// TIA Portal project "Milk_P_2" (V17)

(* hardware
DEVICE "S7-1200 station_1"  S7-1200 Station
   slot 0: "Rack_0"  S7-1200 Rack  Rack  V1.0
   slot 1: "PLC_1"  CPU 1217C DC/DC/DC  6ES7 217-1AG40-0XB0  V4.5
   slot 2: "DI 8x24VDC_1"  6ES7 221-1BF32-0XB0  V2.0
   slot 3: "DQ 8x24VDC _1"  SM 1222 DQ8 x 24VDC  6ES7 222-1BF32-0XB0  V2.0
DEVICE "HMI_1"  KTP700 Basic PN
   slot 0: "HMI_1"  KTP700 Basic PN  6AV2 123-2GB03-0AX0  17.0.0.0
   slot 1: "HMI_RT_1"  KTP700 Basic PN  6AV2 123-2GB03-0AX0  17.0.0.0
   slot 5: "HMI_1.IE_CP_1"  PROFINET Interface  17.0.0.0
      slot 1: "PROFINET Interface_1"  PROFINET Interface
         slot 1: "Port_1"  Port
*)

// ===== PLC "PLC_1"  CPU 1217C DC/DC/DC =====

VAR_GLOBAL   // PLC tag table "Default tag table"
   "Cycle_on_Memory_Bit" AT %M100.0 : Bool;
   "Low_Level_Sensor" AT %M1.0 : Bool;
   "High_Level_Sensor" AT %M1.1 : Bool;
   "Pump_1" AT %Q1.0 : Bool;
   "Milk_Level" AT %MD50 : Real;
   "Start_Fill" AT %M2.0 : Bool;
   "Stop_Fill" AT %M2.1 : Bool;
   "Drain_Start" AT %M2.2 : Bool;
   "Drain_Stop" AT %M2.3 : Bool;
   "Cycle_on_Memory_Bit_2" AT %M200.0 : Bool;
   "Pump_2" AT %Q1.1 : Bool;
   "Sep_Start" AT %M2.4 : Bool;
   "Sep_Stop" AT %M2.5 : Bool;
   "Sep_Memory_Bit" AT %M2.6 : Bool;
   "Clock_Byte" AT %MB0 : Byte;
   "Clock_10Hz" AT %M0.0 : Bool;
   "Clock_5Hz" AT %M0.1 : Bool;
   "Clock_2.5Hz" AT %M0.2 : Bool;
   "Clock_2Hz" AT %M0.3 : Bool;
   "Clock_1.25Hz" AT %M0.4 : Bool;
   "Clock_1Hz" AT %M0.5 : Bool;
   "Clock_0.625Hz" AT %M0.6 : Bool;
   "Clock_0.5Hz" AT %M0.7 : Bool;
   "HMI_Mixer" AT %M2.7 : Bool;
   "Pump_3" AT %Q0.3 : Bool;
   "Furnace_ON" AT %M4.3 : Bool;
   "Furnace_Temp_Sensor" AT %MW4 : Int;
   "Cycle_on_Memory_Bit_3" AT %M50.0 : Bool;
   "Current_Milk_Temp" AT %MW8 : Int;
   "Start_HE" AT %M1.2 : Bool;
   "Stop_HE" AT %M1.3 : Bool;
   "memory_1" AT %M1.4 : Bool;
   "Inıtial_Milk_Temp" AT %MW16 : Int;
   "Wanted_Milk_Temp" AT %MW10 : Int;
   "Heating" AT %Q0.4 : Bool;
   "Cooling_Temp_Sensor" AT %MW12 : Int;
   "Cooling_ON" AT %M1.5 : Bool;
   "Start_CL" AT %M1.6 : Bool;
   "Stop_CL" AT %M1.7 : Bool;
   "Cycle_on_Memory_Bit_4" AT %M7.0 : Bool;
   "memory_2" AT %M7.1 : Bool;
   "Cold_Milk_Temp" AT %MW14 : Int;
   "Heating_OFF" AT %M7.2 : Bool;
   "Cooling_OFF" AT %M7.4 : Bool;
   "Milk_Level_2" AT %MD18 : Real;
   "Low_Level_2" AT %M22.0 : Bool;
   "High_Level_2" AT %M26.0 : Bool;
   "Memory_3" AT %M7.5 : Bool;
   "working" AT %M28.0 : Bool;
   "Start_Package" AT %M28.1 : Bool;
END_VAR

DATA_BLOCK "Bottle Calculation_DB"   // DB1
{ S7_Optimized_Access := 'TRUE' }
VERSION : 0.1
// stored: InstanceOfName Bottle Calculation
"Bottle Calculation"
BEGIN
END_DATA_BLOCK

DATA_BLOCK "Cooling_DB"   // DB2
{ S7_Optimized_Access := 'TRUE' }
VERSION : 0.1
// stored: InstanceOfName Cooling
"Cooling"
BEGIN
END_DATA_BLOCK

DATA_BLOCK "Milk_Pasteurization_DB"   // DB9
{ S7_Optimized_Access := 'TRUE' }
VERSION : 0.1
   VAR
      Fire_Alarm : Bool;
      Warning_Lights : Bool;
      Water_Mist_System : Bool;
   END_VAR
BEGIN
END_DATA_BLOCK

DATA_BLOCK "Heat_Exchange_DB_1"   // DB11
{ S7_Optimized_Access := 'TRUE' }
VERSION : 0.1
// stored: InstanceOfName Heat_Exchange
"Heat_Exchange"
BEGIN
END_DATA_BLOCK

DATA_BLOCK "Pasteurized_Tank_fill_DB"   // DB12
{ S7_Optimized_Access := 'TRUE' }
VERSION : 0.1
// stored: InstanceOfName Pasteurized_Tank_fill
"Pasteurized_Tank_fill"
BEGIN
END_DATA_BLOCK

DATA_BLOCK "Tank_Fill_Drain_DB_1"   // DB13
{ S7_Optimized_Access := 'TRUE' }
VERSION : 0.1
// stored: InstanceOfName Tank_Fill_Drain
"Tank_Fill_Drain"
BEGIN
END_DATA_BLOCK

DATA_BLOCK "Fat_Seperator_DB"   // DB14
{ S7_Optimized_Access := 'TRUE' }
VERSION : 0.1
// stored: InstanceOfName Fat_Seperator
"Fat_Seperator"
BEGIN
END_DATA_BLOCK

// folder: System blocks/Program resources

DATA_BLOCK "Milk_Tank_Timer_1"   // DB3
{ S7_Optimized_Access := 'TRUE' }
AUTHOR : Simatic
FAMILY : IEC
NAME : IEC_TMR
VERSION : 1.0
// stored: InstanceOfName IEC_TIMER
"IEC_TIMER"
BEGIN
END_DATA_BLOCK

DATA_BLOCK "Milk_Tank_Timer_2"   // DB4
{ S7_Optimized_Access := 'TRUE' }
AUTHOR : Simatic
FAMILY : IEC
NAME : IEC_TMR
VERSION : 1.0
// stored: InstanceOfName IEC_TIMER
"IEC_TIMER"
BEGIN
END_DATA_BLOCK

DATA_BLOCK "Sep_Timer"   // DB5
{ S7_Optimized_Access := 'TRUE' }
AUTHOR : Simatic
FAMILY : IEC
NAME : IEC_TMR
VERSION : 1.0
// stored: InstanceOfName IEC_TIMER
"IEC_TIMER"
BEGIN
END_DATA_BLOCK

DATA_BLOCK "HE_Timer1"   // DB6
{ S7_Optimized_Access := 'TRUE' }
AUTHOR : Simatic
FAMILY : IEC
NAME : IEC_TMR
VERSION : 1.0
// stored: InstanceOfName IEC_TIMER
"IEC_TIMER"
BEGIN
END_DATA_BLOCK

DATA_BLOCK "Cooling_Timer"   // DB7
{ S7_Optimized_Access := 'TRUE' }
AUTHOR : Simatic
FAMILY : IEC
NAME : IEC_TMR
VERSION : 1.0
// stored: InstanceOfName IEC_TIMER
"IEC_TIMER"
BEGIN
END_DATA_BLOCK

DATA_BLOCK "P_Tank_Timer1"   // DB8
{ S7_Optimized_Access := 'TRUE' }
AUTHOR : Simatic
FAMILY : IEC
NAME : IEC_TMR
VERSION : 1.0
// stored: InstanceOfName IEC_TIMER
"IEC_TIMER"
BEGIN
END_DATA_BLOCK

DATA_BLOCK "Bottle Counter"   // DB10
{ S7_Optimized_Access := 'TRUE' }
AUTHOR : Simatic
FAMILY : IEC
NAME : CNTR
VERSION : 1.0
// stored: InstanceOfName IEC_COUNTER
"IEC_COUNTER"
BEGIN
END_DATA_BLOCK

// folder: (top level)

FUNCTION_BLOCK "Tank_Fill_Drain"   // FB1, LAD
{ S7_Optimized_Access := 'TRUE' }
VERSION : 0.1
   VAR_INPUT
      "Fill Start" : Bool;
      "Fill Stop" : Bool;
      "Drain Start" : Bool;
      "Drain Stop" : Bool;
   END_VAR
   VAR_OUTPUT
      "Milk Level" : Real;
      "Low Level" : Bool;
      "Pump 2" : Bool;
      Pump : Bool;
      "High Level" : Bool;
   END_VAR
   VAR
      Inıtial_Fat_P : Real := 4.0;
   END_VAR
   VAR_TEMP
      Fat_temp : Real;
   END_VAR
   VAR_TEMP   // added for the SCL form of the ladder/FBD networks
      _w1 : Bool;
   END_VAR
BEGIN

REGION Network 1: Start_Fill System
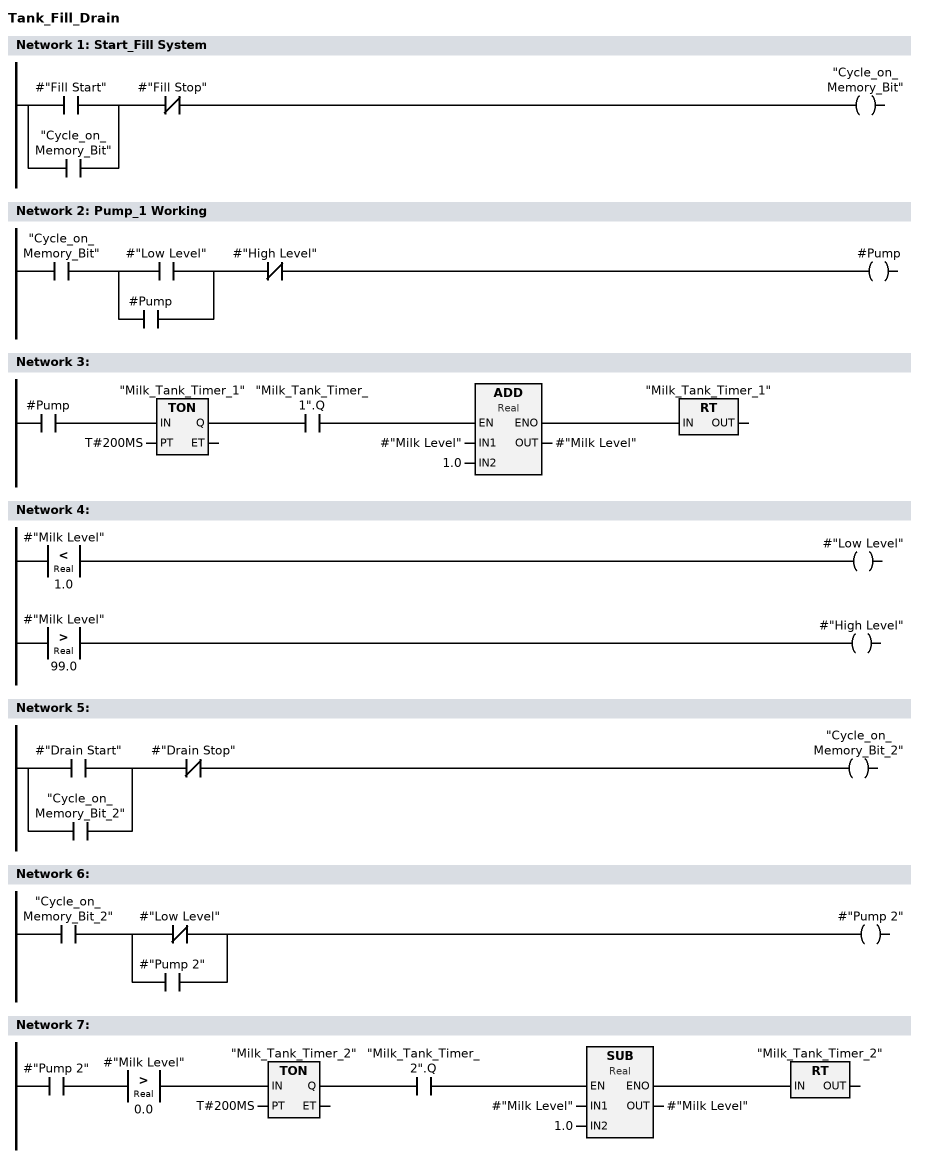
   RUNG wire#powerrail
      Contact( #"Fill Start" )
      wire#w1
      I_Contact( #"Fill Stop" )
      Coil( "Cycle_on_Memory_Bit" )
   END_RUNG
   RUNG wire#powerrail
      Contact( "Cycle_on_Memory_Bit" )
   END_RUNG wire#w1
   // the same network as SCL:
   "Cycle_on_Memory_Bit" := (#"Fill Start" OR "Cycle_on_Memory_Bit") AND NOT #"Fill Stop";
END_REGION

REGION Network 2: Pump_1 Working
   RUNG wire#powerrail
      Contact( "Cycle_on_Memory_Bit" )
      wire#w1
      Contact( #"Low Level" )
      wire#w2
      I_Contact( #"High Level" )
      Coil( #Pump )
   END_RUNG
   RUNG wire#w1
      Contact( #Pump )
   END_RUNG wire#w2
   // the same network as SCL:
   #Pump := "Cycle_on_Memory_Bit" AND (#"Low Level" OR #Pump) AND NOT #"High Level";
END_REGION

REGION Network 3
   "Milk_Tank_Timer_1".TON(IN := #Pump, PT := T#200MS);
   #_w1 := "Milk_Tank_Timer_1".Q AND "Milk_Tank_Timer_1".Q;
   IF #_w1 THEN
       #"Milk Level" := #"Milk Level" + 1.0;
       RESET_TIMER("Milk_Tank_Timer_1");
   END_IF;
END_REGION

REGION Network 4
   RUNG wire#powerrail
      { S7_Templates := "SrcType := Real" } LT_Contact(in1 := #"Milk Level", in2 := 1.0)
      Coil( #"Low Level" )
   END_RUNG
   RUNG wire#powerrail
      { S7_Templates := "SrcType := Real" } GT_Contact(in1 := #"Milk Level", in2 := 99.0)
      Coil( #"High Level" )
   END_RUNG
   // the same network as SCL:
   #"Low Level" := #"Milk Level" < 1.0;
   #"High Level" := #"Milk Level" > 99.0;
END_REGION

REGION Network 5
   RUNG wire#powerrail
      Contact( #"Drain Start" )
      wire#w1
      I_Contact( #"Drain Stop" )
      Coil( "Cycle_on_Memory_Bit_2" )
   END_RUNG
   RUNG wire#powerrail
      Contact( "Cycle_on_Memory_Bit_2" )
   END_RUNG wire#w1
   // the same network as SCL:
   "Cycle_on_Memory_Bit_2" := (#"Drain Start" OR "Cycle_on_Memory_Bit_2") AND NOT #"Drain Stop";
END_REGION

REGION Network 6
   RUNG wire#powerrail
      Contact( "Cycle_on_Memory_Bit_2" )
      wire#w1
      I_Contact( #"Low Level" )
      wire#w2
      Coil( #"Pump 2" )
   END_RUNG
   RUNG wire#w1
      Contact( #"Pump 2" )
   END_RUNG wire#w2
   // the same network as SCL:
   #"Pump 2" := "Cycle_on_Memory_Bit_2" AND (NOT #"Low Level" OR #"Pump 2");
END_REGION

REGION Network 7
   "Milk_Tank_Timer_2".TON(IN := #"Pump 2" AND (#"Milk Level" > 0.0), PT := T#200MS);
   #_w1 := "Milk_Tank_Timer_2".Q AND "Milk_Tank_Timer_2".Q;
   IF #_w1 THEN
       #"Milk Level" := #"Milk Level" - 1.0;
       RESET_TIMER("Milk_Tank_Timer_2");
   END_IF;
END_REGION
END_FUNCTION_BLOCK

FUNCTION_BLOCK "Heat_Exchange"   // FB2, LAD
{ S7_Optimized_Access := 'TRUE' }
VERSION : 0.1
   VAR_INPUT
      "Heat Exchanger Start" : Bool;
      "Heat Exchanger Stop" : Bool;
   END_VAR
   VAR_OUTPUT
      "Furnace ON" : Bool;
      "Current Milk Temperature" : Int;
   END_VAR
   VAR
      heat_difference : Int;
      addition_step : Int;
      furnace_temp_sensor : Int := 500;
      "wanted milk temp" : Int := 72;
      "Initial Temperature" : Int := 20;
   END_VAR
   VAR_TEMP   // added for the SCL form of the ladder/FBD networks
      _w1 : Bool;
   END_VAR
BEGIN

REGION Network 1
   // While loop
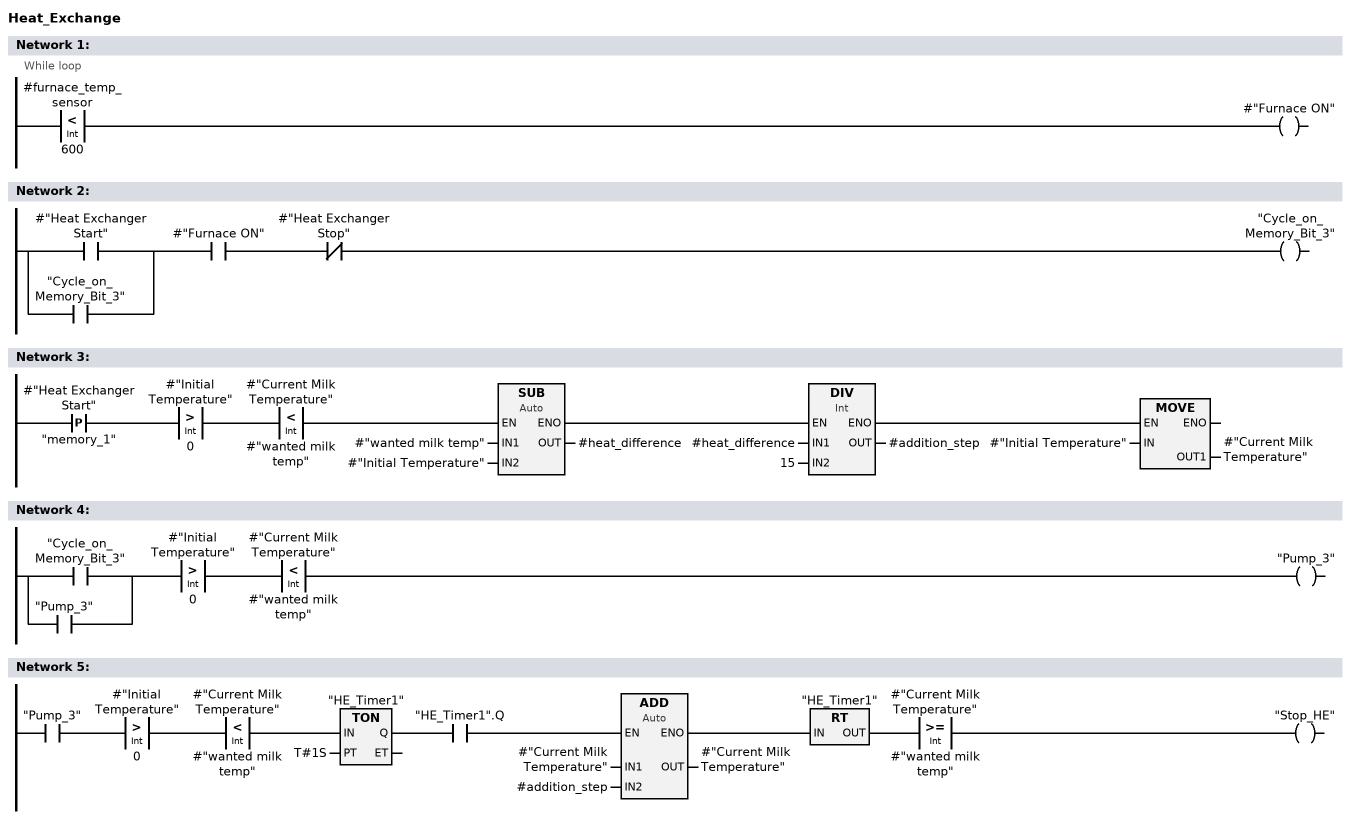
   RUNG wire#powerrail
      { S7_Templates := "SrcType := Int" } LT_Contact(in1 := #furnace_temp_sensor, in2 := 600)
      Coil( #"Furnace ON" )
   END_RUNG
   // the same network as SCL:
   #"Furnace ON" := #furnace_temp_sensor < 600;
END_REGION

REGION Network 2
   RUNG wire#powerrail
      Contact( #"Heat Exchanger Start" )
      wire#w1
      Contact( #"Furnace ON" )
      I_Contact( #"Heat Exchanger Stop" )
      Coil( "Cycle_on_Memory_Bit_3" )
   END_RUNG
   RUNG wire#powerrail
      Contact( "Cycle_on_Memory_Bit_3" )
   END_RUNG wire#w1
   // the same network as SCL:
   "Cycle_on_Memory_Bit_3" := (#"Heat Exchanger Start" OR "Cycle_on_Memory_Bit_3") AND #"Furnace ON" AND NOT #"Heat Exchanger Stop";
END_REGION

REGION Network 3
   RUNG wire#powerrail
      P_Contact(operand := #"Heat Exchanger Start", bit := "memory_1")
      { S7_Templates := "SrcType := Int" } GT_Contact(in1 := #"Initial Temperature", in2 := 0)
      { S7_Templates := "SrcType := Int" } LT_Contact(in1 := #"Current Milk Temperature", in2 := #"wanted milk temp")
      Sub(in1 := #"wanted milk temp", in2 := #"Initial Temperature", out => #heat_difference)
      { S7_Templates := "SrcType := Int" } Div(in1 := #heat_difference, in2 := 15, out => #addition_step)
      Move(in := #"Initial Temperature", out1 => #"Current Milk Temperature")
   END_RUNG
   // the same network as SCL:
   #_w1 := #"Heat Exchanger Start" AND NOT "memory_1";   // rising edge of #"Heat Exchanger Start"
   "memory_1" := #"Heat Exchanger Start";
   IF #_w1 AND (#"Initial Temperature" > 0) AND (#"Current Milk Temperature" < #"wanted milk temp") THEN
       #heat_difference := #"wanted milk temp" - #"Initial Temperature";
       #addition_step := #heat_difference / 15;
       #"Current Milk Temperature" := #"Initial Temperature";
   END_IF;
END_REGION

REGION Network 4
   RUNG wire#powerrail
      Contact( "Cycle_on_Memory_Bit_3" )
      wire#w1
      { S7_Templates := "SrcType := Int" } GT_Contact(in1 := #"Initial Temperature", in2 := 0)
      { S7_Templates := "SrcType := Int" } LT_Contact(in1 := #"Current Milk Temperature", in2 := #"wanted milk temp")
      Coil( "Pump_3" )
   END_RUNG
   RUNG wire#powerrail
      Contact( "Pump_3" )
   END_RUNG wire#w1
   // the same network as SCL:
   "Pump_3" := ("Cycle_on_Memory_Bit_3" OR "Pump_3") AND (#"Initial Temperature" > 0) AND (#"Current Milk Temperature" < #"wanted milk temp");
END_REGION

REGION Network 5
   "HE_Timer1".TON(IN := "Pump_3" AND (#"Initial Temperature" > 0) AND (#"Current Milk Temperature" < #"wanted milk temp"),
                   PT := T#1S);
   #_w1 := "HE_Timer1".Q AND "HE_Timer1".Q;
   IF #_w1 THEN
       #"Current Milk Temperature" := #"Current Milk Temperature" + #addition_step;
       RESET_TIMER("HE_Timer1");
   END_IF;
   "Stop_HE" := #_w1 AND (#"Current Milk Temperature" >= #"wanted milk temp");
END_REGION
END_FUNCTION_BLOCK

FUNCTION_BLOCK "Cooling"   // FB3, LAD
{ S7_Optimized_Access := 'TRUE' }
VERSION : 0.1
   VAR_OUTPUT
      "Cooling OFF" : Bool;
      "Cooling ON" : Bool;
   END_VAR
   VAR
      heat_diff : Int;
      diff_step : Int;
      Wanted_cold_milk : Int := 4;
      "Current Temp" : Int;
      cooling_temp_sensor : Int := -15;
   END_VAR
   VAR_TEMP   // added for the SCL form of the ladder/FBD networks
      _w1 : Bool;
   END_VAR
BEGIN

REGION Network 1
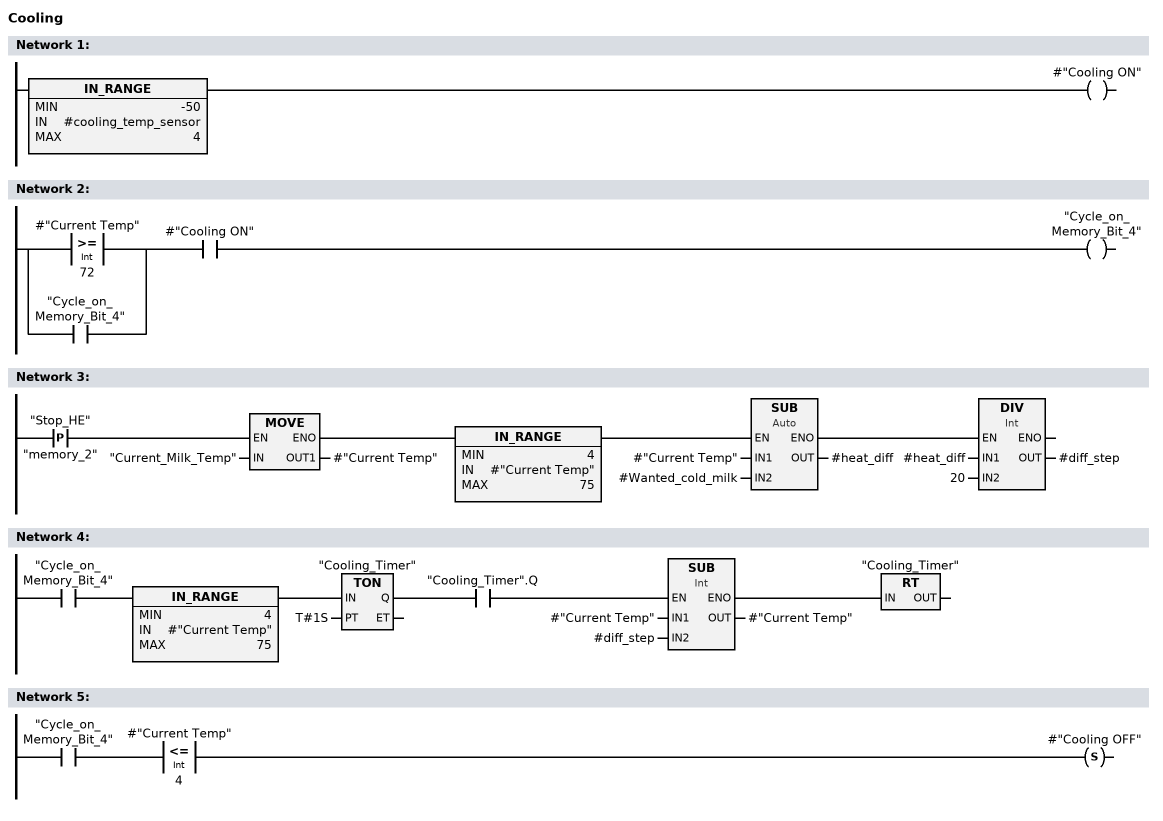
   RUNG wire#powerrail
      { S7_Templates := "SrcType := Int" } InRange(min := -50, in := #cooling_temp_sensor, max := 4)
      Coil( #"Cooling ON" )
   END_RUNG
   // the same network as SCL:
   #"Cooling ON" := (-50 <= #cooling_temp_sensor) AND (#cooling_temp_sensor <= 4);
END_REGION

REGION Network 2
   RUNG wire#powerrail
      { S7_Templates := "SrcType := Int" } GE_Contact(in1 := #"Current Temp", in2 := 72)
      wire#w1
      Contact( #"Cooling ON" )
      Coil( "Cycle_on_Memory_Bit_4" )
   END_RUNG
   RUNG wire#powerrail
      Contact( "Cycle_on_Memory_Bit_4" )
   END_RUNG wire#w1
   // the same network as SCL:
   "Cycle_on_Memory_Bit_4" := ((#"Current Temp" >= 72) OR "Cycle_on_Memory_Bit_4") AND #"Cooling ON";
END_REGION

REGION Network 3
   RUNG wire#powerrail
      P_Contact(operand := "Stop_HE", bit := "memory_2")
      Move(in := "Current_Milk_Temp", out1 => #"Current Temp")
      { S7_Templates := "SrcType := Int" } InRange(min := 4, in := #"Current Temp", max := 75)
      Sub(in1 := #"Current Temp", in2 := #Wanted_cold_milk, out => #heat_diff)
      { S7_Templates := "SrcType := Int" } Div(in1 := #heat_diff, in2 := 20, out => #diff_step)
   END_RUNG
   // the same network as SCL:
   #_w1 := "Stop_HE" AND NOT "memory_2";   // rising edge of "Stop_HE"
   "memory_2" := "Stop_HE";
   IF #_w1 THEN #"Current Temp" := "Current_Milk_Temp"; END_IF;
   IF #_w1 AND (4 <= #"Current Temp") AND (#"Current Temp" <= 75) THEN
       #heat_diff := #"Current Temp" - #Wanted_cold_milk;
       #diff_step := #heat_diff / 20;
   END_IF;
END_REGION

REGION Network 4
   "Cooling_Timer".TON(IN := "Cycle_on_Memory_Bit_4" AND (4 <= #"Current Temp") AND (#"Current Temp" <= 75),
                       PT := T#1S);
   #_w1 := "Cooling_Timer".Q AND "Cooling_Timer".Q;
   IF #_w1 THEN
       #"Current Temp" := #"Current Temp" - #diff_step;
       RESET_TIMER("Cooling_Timer");
   END_IF;
END_REGION

REGION Network 5
   RUNG wire#powerrail
      Contact( "Cycle_on_Memory_Bit_4" )
      { S7_Templates := "SrcType := Int" } LE_Contact(in1 := #"Current Temp", in2 := 4)
      S_Coil( #"Cooling OFF" )
   END_RUNG
   // the same network as SCL:
   IF "Cycle_on_Memory_Bit_4" AND (#"Current Temp" <= 4) THEN #"Cooling OFF" := TRUE; END_IF;
END_REGION
END_FUNCTION_BLOCK

FUNCTION_BLOCK "Fat_Seperator"   // FB4, LAD
{ S7_Optimized_Access := 'TRUE' }
VERSION : 0.1
   VAR_INPUT
      "Seperator Start" : Bool;
      "Seperator Stop" : Bool;
   END_VAR
   VAR_OUTPUT
      "Fat Percantage" : Int := 4;
   END_VAR
   VAR
      wanted_fat : Int := 2;
      diff : Int;
   END_VAR
BEGIN

REGION Network 1
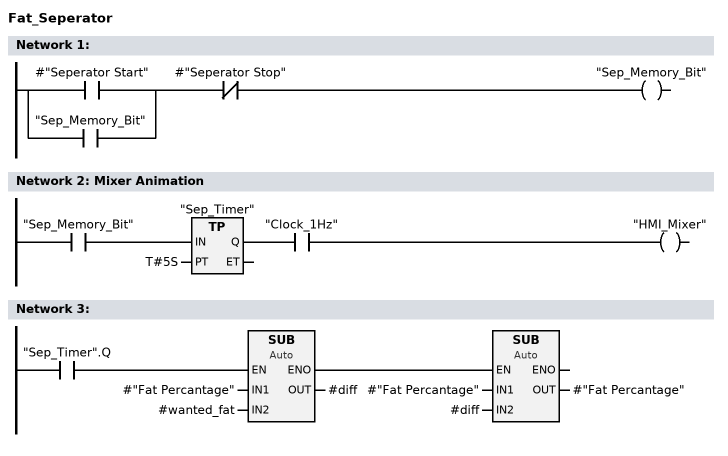
   RUNG wire#powerrail
      Contact( #"Seperator Start" )
      wire#w1
      I_Contact( #"Seperator Stop" )
      Coil( "Sep_Memory_Bit" )
   END_RUNG
   RUNG wire#powerrail
      Contact( "Sep_Memory_Bit" )
   END_RUNG wire#w1
   // the same network as SCL:
   "Sep_Memory_Bit" := (#"Seperator Start" OR "Sep_Memory_Bit") AND NOT #"Seperator Stop";
END_REGION

REGION Network 2: Mixer Animation
   "Sep_Timer".TP(IN := "Sep_Memory_Bit", PT := T#5S);
   "HMI_Mixer" := "Sep_Timer".Q AND "Clock_1Hz";
END_REGION

REGION Network 3
   RUNG wire#powerrail
      Contact( "Sep_Timer".Q )
      Sub(in1 := #"Fat Percantage", in2 := #wanted_fat, out => #diff)
      Sub(in1 := #"Fat Percantage", in2 := #diff, out => #"Fat Percantage")
   END_RUNG
   // the same network as SCL:
   IF "Sep_Timer".Q THEN
       #diff := #"Fat Percantage" - #wanted_fat;
       #"Fat Percantage" := #"Fat Percantage" - #diff;
   END_IF;
END_REGION
END_FUNCTION_BLOCK

FUNCTION_BLOCK "Pasteurized_Tank_fill"   // FB5, LAD
{ S7_Optimized_Access := 'TRUE' }
VERSION : 0.1
   VAR_INPUT
      Start : Bool;
      Stop : Bool;
   END_VAR
   VAR_OUTPUT
      low : Bool;
      high : Bool;
      working : Bool;
      milk_level : Real;
   END_VAR
   VAR_TEMP   // added for the SCL form of the ladder/FBD networks
      _w1 : Bool;
   END_VAR
BEGIN

REGION Network 1
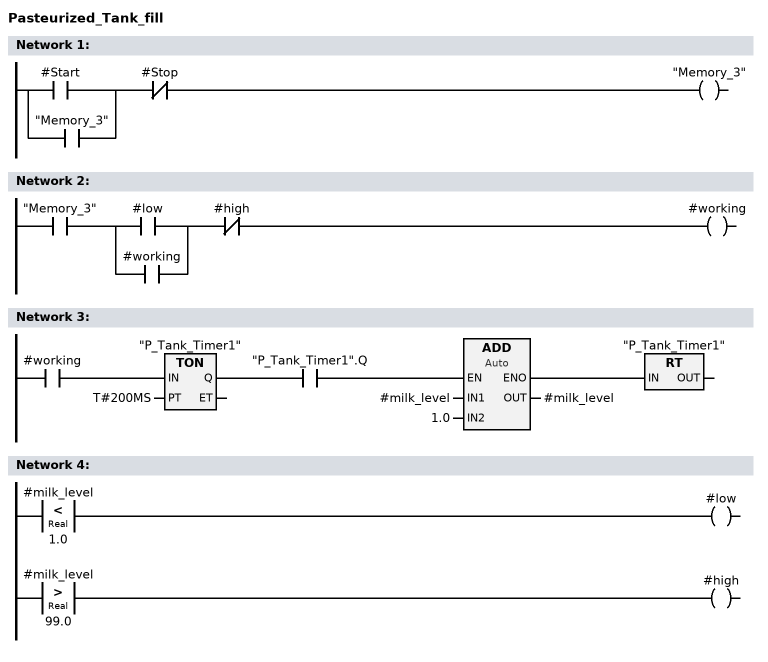
   RUNG wire#powerrail
      Contact( #Start )
      wire#w1
      I_Contact( #Stop )
      Coil( "Memory_3" )
   END_RUNG
   RUNG wire#powerrail
      Contact( "Memory_3" )
   END_RUNG wire#w1
   // the same network as SCL:
   "Memory_3" := (#Start OR "Memory_3") AND NOT #Stop;
END_REGION

REGION Network 2
   RUNG wire#powerrail
      Contact( "Memory_3" )
      wire#w1
      Contact( #low )
      wire#w2
      I_Contact( #high )
      Coil( #working )
   END_RUNG
   RUNG wire#w1
      Contact( #working )
   END_RUNG wire#w2
   // the same network as SCL:
   #working := "Memory_3" AND (#low OR #working) AND NOT #high;
END_REGION

REGION Network 3
   "P_Tank_Timer1".TON(IN := #working, PT := T#200MS);
   #_w1 := "P_Tank_Timer1".Q AND "P_Tank_Timer1".Q;
   IF #_w1 THEN
       #milk_level := #milk_level + 1.0;
       RESET_TIMER("P_Tank_Timer1");
   END_IF;
END_REGION

REGION Network 4
   RUNG wire#powerrail
      { S7_Templates := "SrcType := Real" } LT_Contact(in1 := #milk_level, in2 := 1.0)
      Coil( #low )
   END_RUNG
   RUNG wire#powerrail
      { S7_Templates := "SrcType := Real" } GT_Contact(in1 := #milk_level, in2 := 99.0)
      Coil( #high )
   END_RUNG
   // the same network as SCL:
   #low := #milk_level < 1.0;
   #high := #milk_level > 99.0;
END_REGION
END_FUNCTION_BLOCK

FUNCTION_BLOCK "Bottle Calculation"   // FB6, LAD
{ S7_Optimized_Access := 'TRUE' }
VERSION : 0.1
   VAR_INPUT
      "Start Packaging" : Bool;
   END_VAR
   VAR_OUTPUT
      "Bottle Count" : Int;
   END_VAR
   VAR
      C1 : Bool;
      "Milk Litres" : Real := 10.0;
      "Bottle Litres" : Real := 0.35;
      Running : Bool;
   END_VAR
   VAR_TEMP   // added for the SCL form of the ladder/FBD networks
      _w1 : Bool;
   END_VAR
BEGIN

REGION Network 1
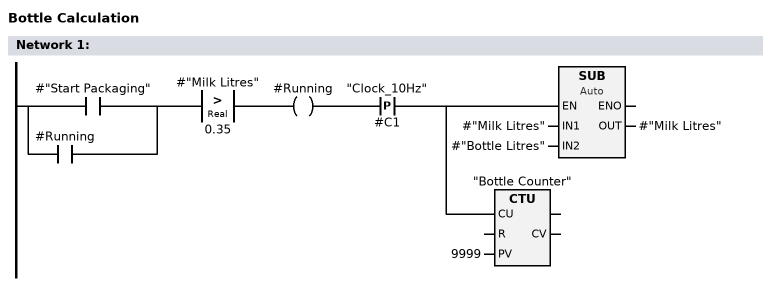
   #Running := (#"Start Packaging" OR #Running) AND (#"Milk Litres" > 0.35);
   #_w1 := #Running AND "Clock_10Hz" AND NOT #C1;   // rising edge of "Clock_10Hz"
   #C1 := "Clock_10Hz";
   IF #_w1 THEN #"Milk Litres" := #"Milk Litres" - #"Bottle Litres"; END_IF;
   "Bottle Counter".CTU(CU := #_w1, PV := 9999);
END_REGION
END_FUNCTION_BLOCK

ORGANIZATION_BLOCK "Main"   // OB1, LAD, ProgramCycle
TITLE = "Main Program Sweep (Cycle)"
{ S7_Optimized_Access := 'TRUE' }
VERSION : 0.1
   VAR_INPUT
      Initial_Call : Bool;   // Initial call of this OB
      Remanence : Bool;   // =True, if remanent data are available
   END_VAR
BEGIN

REGION Network 1: Raw Milk Fill and Drain System
   // Raw milk is filled to a storage tank and it is drain to a fat seperator system.
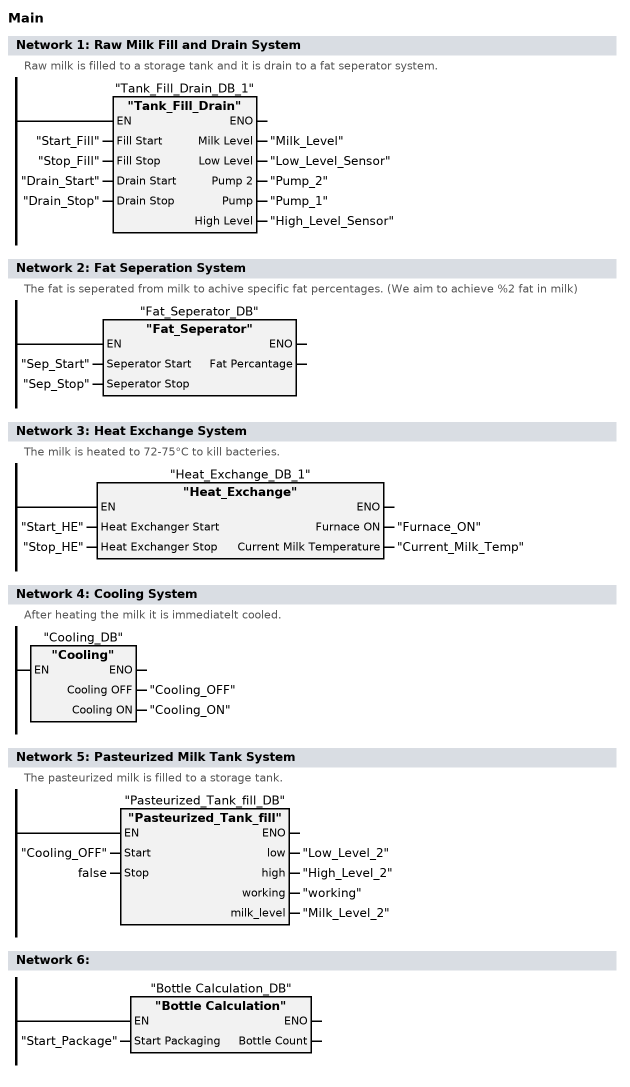
   RUNG wire#powerrail
      "Tank_Fill_Drain_DB_1"("Fill Start" := "Start_Fill", "Fill Stop" := "Stop_Fill", "Drain Start" := "Drain_Start", "Drain Stop" := "Drain_Stop", "Milk Level" => "Milk_Level", "Low Level" => "Low_Level_Sensor", "Pump 2" => "Pump_2", Pump => "Pump_1", "High Level" => "High_Level_Sensor")
   END_RUNG
   // the same network as SCL:
   "Tank_Fill_Drain_DB_1"("Fill Start" := "Start_Fill",   // "Tank_Fill_Drain"
                          "Fill Stop" := "Stop_Fill",
                          "Drain Start" := "Drain_Start",
                          "Drain Stop" := "Drain_Stop",
                          "Milk Level" => "Milk_Level",
                          "Low Level" => "Low_Level_Sensor",
                          "Pump 2" => "Pump_2",
                          Pump => "Pump_1",
                          "High Level" => "High_Level_Sensor");
END_REGION

REGION Network 2: Fat Seperation System
   // The fat is seperated from milk to achive specific fat percentages. (We aim to achieve %2 fat in milk)
   RUNG wire#powerrail
      "Fat_Seperator_DB"("Seperator Start" := "Sep_Start", "Seperator Stop" := "Sep_Stop", "Fat Percantage" =>)
   END_RUNG
   // the same network as SCL:
   "Fat_Seperator_DB"("Seperator Start" := "Sep_Start", "Seperator Stop" := "Sep_Stop");   // "Fat_Seperator"
END_REGION

REGION Network 3: Heat Exchange System
   // The milk is heated to 72-75°C to kill bacteries.
   RUNG wire#powerrail
      "Heat_Exchange_DB_1"("Heat Exchanger Start" := "Start_HE", "Heat Exchanger Stop" := "Stop_HE", "Furnace ON" => "Furnace_ON", "Current Milk Temperature" => "Current_Milk_Temp")
   END_RUNG
   // the same network as SCL:
   "Heat_Exchange_DB_1"("Heat Exchanger Start" := "Start_HE",   // "Heat_Exchange"
                        "Heat Exchanger Stop" := "Stop_HE",
                        "Furnace ON" => "Furnace_ON",
                        "Current Milk Temperature" => "Current_Milk_Temp");
END_REGION

REGION Network 4: Cooling System
   // After heating the milk it is immediatelt cooled.
   RUNG wire#powerrail
      "Cooling_DB"("Cooling OFF" => "Cooling_OFF", "Cooling ON" => "Cooling_ON")
   END_RUNG
   // the same network as SCL:
   "Cooling_DB"("Cooling OFF" => "Cooling_OFF", "Cooling ON" => "Cooling_ON");   // "Cooling"
END_REGION

REGION Network 5: Pasteurized Milk Tank System
   // The pasteurized milk is filled to a storage tank.
   RUNG wire#powerrail
      "Pasteurized_Tank_fill_DB"(Start := "Cooling_OFF", Stop := false, low => "Low_Level_2", high => "High_Level_2", working => "working", milk_level => "Milk_Level_2")
   END_RUNG
   // the same network as SCL:
   "Pasteurized_Tank_fill_DB"(Start := "Cooling_OFF",   // "Pasteurized_Tank_fill"
                           Stop := false,
                           low => "Low_Level_2",
                           high => "High_Level_2",
                           working => "working",
                           milk_level => "Milk_Level_2");
END_REGION

REGION Network 6
   RUNG wire#powerrail
      "Bottle Calculation_DB"("Start Packaging" := "Start_Package", "Bottle Count" =>)
   END_RUNG
   // the same network as SCL:
   "Bottle Calculation_DB"("Start Packaging" := "Start_Package");   // "Bottle Calculation"
END_REGION
END_ORGANIZATION_BLOCK

ORGANIZATION_BLOCK "Cyclic interrupt (HE_FIRE)"   // OB30, LAD, CyclicInterrupt
{ S7_Optimized_Access := 'TRUE' }
VERSION : 0.1
   VAR_INPUT
      Initial_Call : Bool;   // Initial call of this OB
      Event_Count : Int;   // Events discarded
   END_VAR
BEGIN

REGION Network 1
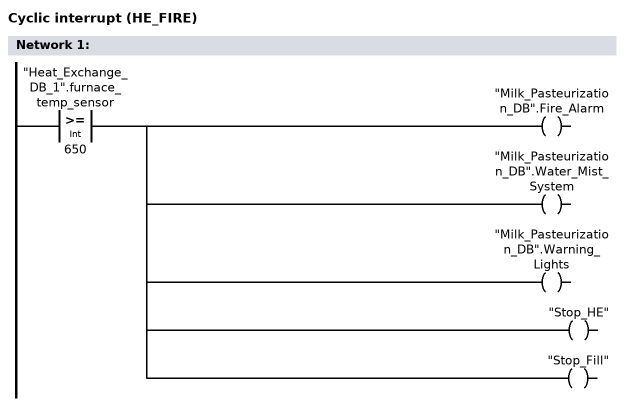
   RUNG wire#powerrail
      { S7_Templates := "SrcType := Int" } GE_Contact(in1 := "Heat_Exchange_DB_1".furnace_temp_sensor, in2 := 650)
      wire#w1
      Coil( "Milk_Pasteurization_DB".Fire_Alarm )
   END_RUNG
   RUNG wire#w1
      Coil( "Milk_Pasteurization_DB".Water_Mist_System )
   END_RUNG
   RUNG wire#w1
      Coil( "Milk_Pasteurization_DB".Warning_Lights )
   END_RUNG
   RUNG wire#w1
      Coil( "Stop_HE" )
   END_RUNG
   RUNG wire#w1
      Coil( "Stop_Fill" )
   END_RUNG
   // the same network as SCL:
   "Milk_Pasteurization_DB".Fire_Alarm := "Heat_Exchange_DB_1".furnace_temp_sensor >= 650;
   "Milk_Pasteurization_DB".Water_Mist_System := "Milk_Pasteurization_DB".Fire_Alarm;
   "Milk_Pasteurization_DB".Warning_Lights := "Milk_Pasteurization_DB".Fire_Alarm;
   "Stop_HE" := "Milk_Pasteurization_DB".Fire_Alarm;
   "Stop_Fill" := "Milk_Pasteurization_DB".Fire_Alarm;
END_REGION
END_ORGANIZATION_BLOCK

(* ===== HMI "HMI_RT_1" =====
system functions are stored by id; their names below are inferred from use
connection "HMI_Connection_1": ETHERNET, SMART_S7_1200_OMS

HMI tags "Default tag table"
   "Tag_ScreenNumber" : UInt, internal
   "Low_Level_Sensor" : Bool = PLC Low_Level_Sensor AT %M1.0, 1 s
   "High_Level_Sensor" : Bool = PLC High_Level_Sensor AT %M1.1, 1 s
   "Water_Level" : Real = PLC Milk_Level AT %MD50, 1 s
   "Start_HMI" : Bool = PLC Start_Fill AT %M2.0, 1 s
   "Stop_HMI" : Bool = PLC Stop_Fill AT %M2.1, 1 s
   "Drain_Start" : Bool = PLC Drain_Start AT %M2.2, 1 s
   "Drain_Stop" : Bool = PLC Drain_Stop AT %M2.3, 1 s
   "Sep_Start" : Bool = PLC Sep_Start AT %M2.4, 100 ms
   "Sep_Stop" : Bool = PLC Sep_Stop AT %M2.5, 100 ms
   "HMI_Mixer" : Bool = PLC HMI_Mixer AT %M2.7, 100 ms
   "Pump_1" : Bool = PLC Pump_1 AT %Q1.0, 100 ms
   "Pump_2" : Bool = PLC Pump_2 AT %Q1.1, 100 ms
   "Start_HE" : Bool = PLC Start_HE AT %M1.2, 1 s
   "Stop_HE" : Bool = PLC Stop_HE AT %M1.3, 1 s
   "Inıtial_Milk_Temp" : Int = PLC Inıtial_Milk_Temp AT %MW16, 1 s
   "Current_Milk_Temp" : Int = PLC Current_Milk_Temp AT %MW8, 1 s
   "Furnace_Temp_Sensor" : Int = PLC Furnace_Temp_Sensor AT %MW4, 1 s
   "Wanted_Milk_Temp" : Int = PLC Wanted_Milk_Temp AT %MW10, 1 s
   "Clock_0.5Hz" : Bool = PLC "Clock_0.5Hz" AT %M0.7, 1 s
   "Clock_10Hz" : Bool = PLC Clock_10Hz AT %M0.0, 1 s
   "Start_CL" : Bool = PLC Start_CL AT %M1.6, 1 s
   "Stop_CL" : Bool = PLC Stop_CL AT %M1.7, 1 s
   "Cold_Milk_Temp" : Int = PLC Cold_Milk_Temp AT %MW14, 1 s
   "Heat_Exchange_DB_1_Initial Temperature" : Int = PLC Heat_Exchange_DB_1."Initial Temperature", 1 s
   "Heat_Exchange_DB_1_wanted milk temp" : Int = PLC Heat_Exchange_DB_1."wanted milk temp", 1 s
   "Heat_Exchange_DB_1_furnace_temp_sensor" : Int = PLC Heat_Exchange_DB_1.furnace_temp_sensor, 1 s
   "Cooling_DB_Wanted_cold_milk" : Int = PLC Cooling_DB.Wanted_cold_milk, 1 s
   "Cooling_DB_Current Temp" : Int = PLC Cooling_DB."Current Temp", 1 s
   "Milk_Level_2" : Real = PLC Milk_Level_2 AT %MD18, 1 s
   "Fat_Seperator_DB_Initial Fat Percantage" : Int = PLC Fat_Seperator_DB."Fat Percantage", 1 s
   "Fat_Seperator_DB_diff" : Int = PLC Fat_Seperator_DB.diff, 1 s
   "Bottle Calculation_DB_Bottle Count" : Int = PLC "Bottle Calculation_DB"."Bottle Count", 1 s
   "Start_Package" : Bool = PLC Start_Package AT %M28.1, 1 s
   "Bottle Counter_CV" : Int = PLC "Bottle Counter".CV, 1 s
   "Low_Level_2" : Bool = PLC Low_Level_2 AT %M22.0, 1 s
   "High_Level_2" : Bool = PLC High_Level_2 AT %M26.0, 1 s

HMI tags "User"
   "Esra Cesur" : WString[254], internal

screen "Root screen" 800x480, template "Template_1"
   on GenerateScreen: SetTag("Stop_HMI", 1)
   Softkey "Softkey_F1" at 0,0 size 0x0
      on KeyDown: ActivateScreen("Root screen", 0)
   Button "Button_3" at 320,349 size 156x119; TextOff 'Cooling'; Authorization "Operator"
      on Click: ActivateScreen("Cooling", 0)
   Button "Button_4" at 479,349 size 156x119; TextOff 'Pasteurized Milk'; Authorization "Operator"
      on Click: ActivateScreen("Pasteurized_Milk", 0)
   Button "Button_5" at 638,349 size 156x119; TextOff 'Log OFF'
      on Click: function_f23ef4c9()
   GraphicView "Graphic view_1" at 0,112 size 800x237; Picture "1009-10099800_cow-milk-cattle"
   Button "Button_2" at 0,349 size 154x119; TextOff 'Raw Milk Tank'; TextOn 'Raw_Milk_Tank'; Authorization "Operator"
      on Click: ActivateScreen("Raw_Milk_Tank", 0)
   Button "Button_1" at 157,349 size 160x119; TextOff 'Heat Exchange'; TextOn 'Heat_Exchange'; Authorization "Operator"
      on Click: ActivateScreen("Heat_Exchange", 0)
   Softkey "Softkey_F8" at 0,0 size 0x0
      on KeyDown: function_f23ef4c9(); ActivateScreen("Root screen", 0)

screen "Raw_Milk_Tank" 800x480
   Softkey "Softkey_F2" at 0,0 size 0x0
      on KeyDown: ActivateScreen("Raw_Milk_Tank", 0)
   Softkey "Softkey_F1" at 0,0 size 0x0
      on KeyDown: ActivateScreen("Root screen", 0)
   GraphicView "Graphic view_19" at 647,214 size 65x49; Picture "Graphic_8"
   GraphicView "Graphic view_18" at 560,291 size 55x48; Picture "Graphic_46"
   GraphicView "Graphic view_10" at 513,97 size 147x222; Picture "Graphic_28"
   GraphicView "Graphic view_12" at 529,133 size 116x119; Picture "Graphic_33"
      Visibility <- "HMI_Mixer"
   GraphicView "Graphic view_11" at 547,126 size 78x94; Picture "Graphic_32"
      Visibility <- "HMI_Mixer"
   GraphicView "Graphic view_20" at 529,133 size 116x119; Picture "Graphic_47"
      Visibility <- "HMI_Mixer"
   GraphicView "Graphic view_21" at 547,126 size 78x94; Picture "Graphic_48"
      Visibility <- "HMI_Mixer"
   GraphicView "Graphic view_23" at 760,215 size 40x51; Picture "Graphic_8"
   GraphicView "Graphic view_17" at 465,140 size 59x47; Picture "Graphic_8"
   GraphicView "Graphic view_7" at 219,338 size 78x57; Picture "Graphic_8"
   GraphicView "Graphic view_3" at 166,340 size 59x53; Picture "Graphic_4"
   GraphicView "Graphic view_1" at 121,113 size 145x239; Picture "Graphic_1"
   Bar "Bar_1" at 138,158 size 112x141; MinimumValue 0; MaximumValue 100
      ProcessValue <- "Water_Level"
   GraphicView "Graphic view_2" at 166,66 size 59x53; Picture "Graphic_3"
   GraphicView "Graphic view_6" at 121,66 size 48x53; Picture "Graphic_8"
   Button "Button_1" at 21,150 size 99x38; TextOff 'Fill Start'
      on Press: function_b14e0dd5("Start_HMI", 0)
      Appearance <- "Start_HMI"
   Button "Button_2" at 21,195 size 100x38; TextOff 'Fill Stop'
      on Press: function_b14e0dd5("Stop_HMI", 0)
      Appearance <- "Stop_HMI"
   Rectangle "Rectangle_1" at 266,253 size 98x22
      Appearance <- "Low_Level_Sensor"
   TextField "Text field_1" at 270,251 size 86x23; Text 'Low Level'
   Rectangle "Rectangle_2" at 266,178 size 101x22
      Appearance <- "High_Level_Sensor"
   TextField "Text field_2" at 270,176 size 90x23; Text 'High Level'
   IOField "I/O field_1" at 151,125 size 88x27; FormatPattern 999
      ProcessValue <- "Water_Level"
   Button "Button_3" at 21,261 size 100x37; TextOff 'Drain Start'
      on Press: function_b14e0dd5("Drain_Start", 0)
      Appearance <- "Drain_Start"
   Button "Button_4" at 21,307 size 100x36; TextOff 'Drain Stop'
      on Press: function_b14e0dd5("Drain_Stop", 0)
      Appearance <- "Drain_Stop"
   GraphicView "Graphic view_5" at 0,66 size 78x53; Picture "Graphic_8"
   GraphicView "Graphic view_4" at 62,70 size 68x46; Picture "Graphic_5"
      Appearance <- "Pump_1"
   GraphicView "Graphic view_9" at 345,337 size 78x57; Picture "Graphic_8"
   GraphicView "Graphic view_8" at 293,345 size 61x45; Picture "Graphic_9"
      Appearance <- "Pump_2"
   GraphicView "Graphic view_14" at 416,339 size 56x54; Picture "Graphic_43"
   GraphicView "Graphic view_15" at 415,174 size 58x170; Picture "Graphic_44"
   GraphicView "Graphic view_16" at 415,139 size 57x48; Picture "Graphic_45"
   TextField "Text field_3" at 534,39 size 97x18; Text 'Fat Percentage'
   Button "Button_5" at 688,347 size 102x35; TextOff 'Mixer Start'
      on Release: ResetBit("Sep_Start")
      on Press: SetBit("Sep_Start")
      Appearance <- "Sep_Start"
   Button "Button_6" at 688,390 size 102x35; TextOff 'Mixer Stop'
      on Release: ResetBit("Sep_Stop")
      on Press: function_b14e0dd5("Sep_Stop", 0)
      Appearance <- "Sep_Stop"
   GraphicView "Graphic view_22" at 490,342 size 190x92; Picture "Graphic_54"
   Group "Group" at 513,97 size 199x242; Picture "Graphic_8"
   TextField "Text field_5" at 526,379 size 120x23; Text 'Seperated Fat'
   GraphicView "Graphic view_13" at 698,217 size 74x44; Picture "Graphic_58"
   IOField "I/O field_2" at 550,58 size 71x32; FormatPattern s99
      ProcessValue <- "Fat_Seperator_DB_Initial Fat Percantage"
   TextField "Text field_4" at 527,61 size 24x23; Text '%'
   Softkey "Softkey_F3" at 0,0 size 0x0
      on KeyDown: ActivateScreen("Heat_Exchange", 0)
   Softkey "Softkey_F4" at 0,0 size 0x0
      on KeyDown: ActivateScreen("Cooling", 0)
   Softkey "Softkey_F5" at 0,0 size 0x0
      on KeyDown: ActivateScreen("Pasteurized_Milk", 0)
   Softkey "Softkey_F8" at 0,0 size 0x0
      on KeyDown: function_f23ef4c9()

screen "Heat_Exchange" 800x480
   GraphicView "Graphic view_1" at 112,33 size 56x55; Picture "Graphic_3"
   GraphicView "Graphic view_2" at 111,78 size 56x318; Picture "Graphic_44"
   GraphicView "Graphic view_3" at 112,389 size 56x56; Picture "Graphic_4"
   GraphicView "Graphic view_4" at 192,390 size 56x54; Picture "Graphic_43"
   GraphicView "Graphic view_8" at 165,391 size 31x53; Picture "Graphic_8"
   GraphicView "Graphic view_5" at 191,90 size 57x308; Picture "Graphic_44"
   GraphicView "Graphic view_17" at 190,43 size 59x55; Picture "Graphic_45"
   GraphicView "Graphic view_18" at 244,42 size 52x57; Picture "Graphic_8"
   GraphicView "Graphic view_15" at 242,41 size 51x320; Picture "Graphic_122"
   GraphicView "Graphic view_9" at 146,354 size 59x50; Picture "Graphic_123"
   GraphicView "Graphic view_10" at 191,355 size 56x46; Picture "Graphic_124"
   GraphicView "Graphic view_11" at 243,355 size 49x47; Picture "Graphic_125"
   GraphicView "Graphic view_7" at 146,41 size 59x320; Picture "Graphic_122"
   Group "Group_1" at 111,33 size 185x412; Picture "Graphic_3"
   Group "Group_2" at 287,44 size 174x397; Picture "Graphic_3"
   GraphicView "Graphic view_28" at 455,101 size 53x378; Picture "Graphic_44"
   GraphicView "Graphic view_27" at 455,54 size 52x55; Picture "Graphic_3"
   GraphicView "Graphic view_19" at 288,44 size 53x53; Picture "Graphic_3"
   GraphicView "Graphic view_20" at 287,87 size 53x306; Picture "Graphic_44"
   GraphicView "Graphic view_21" at 288,387 size 53x54; Picture "Graphic_4"
   GraphicView "Graphic view_22" at 363,388 size 53x52; Picture "Graphic_43"
   GraphicView "Graphic view_23" at 338,389 size 29x51; Picture "Graphic_8"
   GraphicView "Graphic view_24" at 362,99 size 54x297; Picture "Graphic_44"
   GraphicView "Graphic view_25" at 361,54 size 55x53; Picture "Graphic_45"
   GraphicView "Graphic view_26" at 412,53 size 49x55; Picture "Graphic_8"
   GraphicView "Graphic view_35" at 415,46 size 51x320; Picture "Graphic_122"
   GraphicView "Graphic view_36" at 319,359 size 59x50; Picture "Graphic_123"
   GraphicView "Graphic view_37" at 364,360 size 56x46; Picture "Graphic_124"
   GraphicView "Graphic view_38" at 416,360 size 49x47; Picture "Graphic_125"
   GraphicView "Graphic view_39" at 319,46 size 59x320; Picture "Graphic_122"
   GraphicView "Graphic view_40" at 536,130 size 64x47; Picture "Graphic_124"
   GraphicView "Graphic view_13" at 498,131 size 45x47; Picture "Graphic_123"
   GraphicView "Graphic view_12" at 498,49 size 45x85; Picture "Graphic_122"
   GraphicView "Graphic view_32" at 498,9 size 45x47; Picture "Graphic_121"
   GraphicView "Graphic view_33" at 459,9 size 42x47; Picture "Graphic_124"
   GraphicView "Graphic view_34" at 413,8 size 50x51; Picture "Graphic_126"
   Group "Group_4" at 319,46 size 147x363; Picture "Graphic_122"
   GraphicView "Graphic view_31" at 322,3 size 53x49; Picture "Graphic_121"
   GraphicView "Graphic view_30" at 286,4 size 42x47; Picture "Graphic_124"
   GraphicView "Graphic view_29" at 240,4 size 52x47; Picture "Graphic_126"
   Group "Group" at 146,41 size 147x363; Picture "Graphic_122"
   Group "Group_3" at 146,3 size 454x406; Picture "Graphic_124"
   GraphicView "Graphic view_41" at 146,0 size 59x75; Picture "Graphic_122"
   Softkey "Softkey_F2" at 0,0 size 0x0
      on KeyDown: ActivateScreen("Raw_Milk_Tank", 0)
   Softkey "Softkey_F3" at 0,0 size 0x0
      on KeyDown: ActivateScreen("Heat_Exchange", 0)
   GraphicView "Graphic view_42" at 641,0 size 68x24; Picture "Graphic_122"
   GraphicView "Graphic view_6" at 568,8 size 216x193; Picture "Graphic_95"
   GraphicView "Graphic view_14" at 0,31 size 60x59; Picture "Graphic_8"
   Group "Group_5" at 146,0 size 454x409; Picture "Graphic_124"
   Group "Group_6" at 111,33 size 397x446; Picture "Graphic_3"
   GraphicView "Graphic view_16" at 40,31 size 83x57; Picture "Graphic_119"
   IOField "I/O field_2" at 15,144 size 81x44; FormatPattern s99
      ProcessValue <- "Heat_Exchange_DB_1_Initial Temperature"
   IOField "I/O field_3" at 346,441 size 53x35; FormatPattern s99
      ProcessValue <- "Current_Milk_Temp"
   Button "Button_1" at 15,225 size 96x32; TextOff 'Start'
      on Press: function_b14e0dd5("Start_HE", 0)
      Appearance <- "Start_HE"
   Button "Button_2" at 15,262 size 96x32; TextOff 'Stop'
      on Press: function_b14e0dd5("Stop_HE", 0)
      Appearance <- "Stop_HE"
   TrendView "Trend view_1" at 508,207 size 283x258
   IOField "I/O field_1" at 12,363 size 82x48; FormatPattern s99
      ProcessValue <- "Heat_Exchange_DB_1_wanted milk temp"
   TextField "Text field_1" at 33,102 size 59x23; Text 'Initial'
   TextField "Text field_2" at 3,118 size 112x23; Text 'Temperature'
   TextField "Text field_3" at 12,321 size 93x23; Text 'Set Output'
   TextField "Text field_4" at 3,337 size 112x23; Text 'Temperature'
   TextField "Text field_5" at 158,446 size 179x23; Text 'Current Temperature'
   IOField "I/O field_4" at 641,20 size 70x50; FormatPattern s999
      ProcessValue <- "Heat_Exchange_DB_1_furnace_temp_sensor"
   TextField "Text field_6" at 91,155 size 24x23; Text '°C'
   TextField "Text field_7" at 87,375 size 24x23; Text '°C'
   TextField "Text field_8" at 399,446 size 24x23; Text '°C'
   Softkey "Softkey_F1" at 0,0 size 0x0
      on KeyDown: ActivateScreen("Root screen", 0)
   Softkey "Softkey_F4" at 0,0 size 0x0
      on KeyDown: ActivateScreen("Cooling", 0)
   Softkey "Softkey_F5" at 0,0 size 0x0
      on KeyDown: ActivateScreen("Pasteurized_Milk", 0)
   Softkey "Softkey_F8" at 0,0 size 0x0
      on KeyDown: function_f23ef4c9()

screen "Cooling" 800x480
   GraphicView "Graphic view_14" at 0,31 size 60x59; Picture "Graphic_8"
   Group "Group_5" at 146,0 size 454x409; Picture "Graphic_124"
   Group "Group_6" at 111,33 size 397x446; Picture "Graphic_3"
   GraphicView "Graphic view_16" at 40,31 size 83x57; Picture "Graphic_119"
   TrendView "Trend view_1" at 508,207 size 283x258
   GraphicView "Graphic view_6" at 580,11 size 175x178; Picture "Graphic_156"
   IOField "I/O field_2" at 6,189 size 81x44; FormatPattern s99
      ProcessValue <- "Cooling_DB_Current Temp"
   TextField "Text field_1" at 31,141 size 16x23; Text 'Text'
   TextField "Text field_2" at 0,159 size 112x23; Text 'Temperature'
   IOField "I/O field_1" at 9,304 size 80x48; FormatPattern s99
      ProcessValue <- "Cooling_DB_Wanted_cold_milk"
   TextField "Text field_3" at 13,262 size 93x23; Text 'Set Output'
   TextField "Text field_4" at 0,278 size 112x23; Text 'Temperature'
   TrendView "Trend view_2" at 508,202 size 283x263
   TextField "Text field_6" at 88,199 size 24x23; Text '°C'
   TextField "Text field_5" at 88,319 size 24x23; Text '°C'
   GraphicView "Graphic view_40" at 536,130 size 64x47; Picture "Graphic_124"
   GraphicView "Graphic view_13" at 498,131 size 45x47; Picture "Graphic_123"
   GraphicView "Graphic view_12" at 498,49 size 45x85; Picture "Graphic_122"
   GraphicView "Graphic view_32" at 498,9 size 45x47; Picture "Graphic_121"
   GraphicView "Graphic view_33" at 459,9 size 42x47; Picture "Graphic_124"
   GraphicView "Graphic view_34" at 413,8 size 50x51; Picture "Graphic_126"
   Group "Group_4" at 319,46 size 147x363; Picture "Graphic_122"
   GraphicView "Graphic view_31" at 322,3 size 53x49; Picture "Graphic_121"
   GraphicView "Graphic view_30" at 286,4 size 42x47; Picture "Graphic_124"
   GraphicView "Graphic view_29" at 240,4 size 52x47; Picture "Graphic_126"
   Group "Group" at 146,41 size 147x363; Picture "Graphic_122"
   GraphicView "Graphic view_35" at 415,46 size 51x320; Picture "Graphic_122"
   GraphicView "Graphic view_36" at 319,359 size 59x50; Picture "Graphic_123"
   GraphicView "Graphic view_37" at 364,360 size 56x46; Picture "Graphic_124"
   GraphicView "Graphic view_38" at 416,360 size 49x47; Picture "Graphic_125"
   GraphicView "Graphic view_39" at 319,46 size 59x320; Picture "Graphic_122"
   GraphicView "Graphic view_15" at 242,41 size 51x320; Picture "Graphic_122"
   GraphicView "Graphic view_9" at 146,354 size 59x50; Picture "Graphic_123"
   GraphicView "Graphic view_10" at 191,355 size 56x46; Picture "Graphic_124"
   GraphicView "Graphic view_11" at 243,355 size 49x47; Picture "Graphic_125"
   GraphicView "Graphic view_7" at 146,41 size 59x320; Picture "Graphic_122"
   Group "Group_3" at 146,3 size 454x406; Picture "Graphic_124"
   GraphicView "Graphic view_41" at 146,0 size 59x75; Picture "Graphic_122"
   GraphicView "Graphic view_1" at 112,33 size 56x55; Picture "Graphic_3"
   GraphicView "Graphic view_2" at 111,78 size 56x318; Picture "Graphic_44"
   GraphicView "Graphic view_3" at 112,389 size 56x56; Picture "Graphic_4"
   GraphicView "Graphic view_4" at 192,390 size 56x54; Picture "Graphic_43"
   GraphicView "Graphic view_8" at 165,391 size 31x53; Picture "Graphic_8"
   GraphicView "Graphic view_5" at 191,90 size 57x308; Picture "Graphic_44"
   GraphicView "Graphic view_17" at 190,43 size 59x55; Picture "Graphic_45"
   GraphicView "Graphic view_18" at 244,42 size 52x57; Picture "Graphic_8"
   Group "Group_1" at 111,33 size 185x412; Picture "Graphic_3"
   Group "Group_2" at 287,44 size 174x397; Picture "Graphic_3"
   GraphicView "Graphic view_28" at 455,101 size 53x378; Picture "Graphic_44"
   GraphicView "Graphic view_27" at 455,54 size 52x55; Picture "Graphic_3"
   GraphicView "Graphic view_19" at 288,44 size 53x53; Picture "Graphic_3"
   GraphicView "Graphic view_20" at 287,87 size 53x306; Picture "Graphic_44"
   GraphicView "Graphic view_21" at 288,387 size 53x54; Picture "Graphic_4"
   GraphicView "Graphic view_22" at 363,388 size 53x52; Picture "Graphic_43"
   GraphicView "Graphic view_23" at 338,389 size 29x51; Picture "Graphic_8"
   GraphicView "Graphic view_24" at 362,99 size 54x297; Picture "Graphic_44"
   GraphicView "Graphic view_25" at 361,54 size 55x53; Picture "Graphic_45"
   GraphicView "Graphic view_26" at 412,53 size 49x55; Picture "Graphic_8"
   Softkey "Softkey_F1" at 0,0 size 0x0
      on KeyDown: ActivateScreen("Root screen", 0)
   Softkey "Softkey_F2" at 0,0 size 0x0
      on KeyDown: ActivateScreen("Raw_Milk_Tank", 0)
   Softkey "Softkey_F3" at 0,0 size 0x0
      on KeyDown: ActivateScreen("Heat_Exchange", 0)
   Softkey "Softkey_F4" at 0,0 size 0x0
      on KeyDown: ActivateScreen("Cooling", 0)
   Softkey "Softkey_F5" at 0,0 size 0x0
      on KeyDown: ActivateScreen("Pasteurized_Milk", 0)
   Softkey "Softkey_F8" at 0,0 size 0x0
      on KeyDown: function_f23ef4c9()

screen "Pasteurized_Milk" 800x480
   Softkey "Softkey_F1" at 0,0 size 0x0
      on KeyDown: ActivateScreen("Root screen", 0)
   Softkey "Softkey_F2" at 0,0 size 0x0
      on KeyDown: ActivateScreen("Raw_Milk_Tank", 0)
   Softkey "Softkey_F3" at 0,0 size 0x0
      on KeyDown: ActivateScreen("Heat_Exchange", 0)
   Softkey "Softkey_F4" at 0,0 size 0x0
      on KeyDown: ActivateScreen("Cooling", 0)
   Softkey "Softkey_F5" at 0,0 size 0x0
      on KeyDown: ActivateScreen("Pasteurized_Milk", 0)
   GraphicView "Graphic view_2" at 381,45 size 75x75; Picture "Graphic_45"
   GraphicView "Graphic view_7" at 449,45 size 350x78; Picture "Graphic_8"
   GraphicView "Graphic view_1" at 305,107 size 241x289; Picture "Graphic_1"
   TextField "Text field_1" at 355,125 size 141x23; Text 'Pasteurized Milk'
   GraphicView "Graphic view_4" at 316,330 size 223x93; Picture "Graphic_162"
   Bar "Bar_1" at 330,163 size 197x171; MinimumValue 0; MaximumValue 100
      ProcessValue <- "Milk_Level_2"
   Button "Button_1" at 100,182 size 96x32; TextOff 'Bottle'
      Appearance <- "Start_Package"
      on Press: SetBit("Start_Package")
   IOField "I/O field_1" at 107,226 size 89x61; FormatPattern s99999
      ProcessValue <- "Bottle Counter_CV"
   TextField "Text field_2" at 66,287 size 205x23; Text 'Produced Bottle Number'
   Rectangle "Rectangle_1" at 553,301 size 98x22
      Appearance <- "Low_Level_2"
   TextField "Text field_3" at 557,299 size 86x23; Text 'Low Level'
   Rectangle "Rectangle_2" at 549,188 size 101x22
      Appearance <- "High_Level_2"
   TextField "Text field_4" at 553,186 size 90x23; Text 'High Level'
   Softkey "Softkey_F8" at 0,0 size 0x0
      on KeyDown: function_f23ef4c9()

scheduled task "Get User Name"
   on Action: function_f41c6f6c("Esra Cesur")
*)